
                                 // Set value with follow val from above 
                                 #tempReturnVal := "LKinLang_SetValue"(parameterValue := #tempParameterValue,
                                                                       parameterPriority := #statParameterDefinition.priorities.valueFlags.remainingDistance,
                                                                       validCountOfParameter := #statValidCounts.valueFlags.remainingDistance,
                                                                       parameterValueMin := #MINVAL_LREAL,
                                                                       parameterValueMax := #MAXVAL_LREAL,
                                                                       properties := #statParameterDefinition.properties,
                                                                       errorString => #statErrorString,
                                                                       parameterCounter := #statElementCounter.valueFlags.remainingDistance,
                                                                       priorityCounter := #statActualCommand.priority.valueFlags[#statActualValueFlagNumber].remainingDistance,
                                                                       modalCMDPrio := #statModalCommand.priority.valueFlags[#statActualValueFlagNumber].remainingDistance,
                                                                       modalPRGPrio := #statModalProgram.priority.valueFlags[#statActualValueFlagNumber].remainingDistance,
                                                                       parameterCounterInLine := #statElementCounterInLine.valueFlags.remainingDistance,
                                                                       pathDataValue := #statPathDataValue,
                                                                       modalCMDPathDataValue := #statModalCmdValue,
                                                                       modalPRGPathDataValue := #statModalPrgValue);

                                 IF #tempReturnVal = 0 THEN // Parameter is ok
                                   #statActualCommand.pathDataElement.valueFlags[#statActualValueFlagNumber].remainingDistance := #statPathDataValue.valueLReal;
                                   #statModalCommand.pathDataElement.valueFlags[#statActualValueFlagNumber].remainingDistance := #statModalCmdValue.valueLReal;
                                   #statModalProgram.pathDataElement.valueFlags[#statActualValueFlagNumber].remainingDistance := #statModalPrgValue.valueLReal;
                                 ELSE
                                   // Error
                                   #statStatus := #ERR_PARSING;
                                   #statErrorString := CONCAT(IN1 := #statErrorString, IN2 := '; Line: ');
                                   #statErrorString := CONCAT(IN1 := #statErrorString, IN2 := UDINT_TO_STRING(#statTokenizedLine.lineNo));
                                   EXIT;
                                 END_IF;
                               END_IF;

                             END_FOR;
                           END_REGION LREAL_FLAGS

                           // Exit loop in case of error
                           IF #statStatus.%X15 THEN
                             EXIT;
                           END_IF;

                         END_IF;
                       END_REGION SET_VALUES_IN_PATH_DATA_ELEMENT

                     END_FOR;

                     // Exit loop in case of error
                     IF #statStatus.%X15 THEN
                       EXIT;
                     END_IF;

                     // Check if right side of equation; if not reset it 
                     IF #statRightSideOfEquation THEN
                       ;
                     ELSE
                       #statRightSideOfEquation := TRUE;
                       #statStringExpression := '';
                     END_IF;

                     // Go to next state
                     #statStateIntern := #STATE_TOKEN_PROCESSED;

                   END_IF;
                 END_REGION TOKEN_IS_PARAMETER

                 // ------------------------------------------------------------------------------------------
                 // Is token variable
                 // Check if token is a defined variable or interface variable
                 // YES: Go to TOKEN_IS_VARIABLE
                 // NO: Go to TOKEN_IS_UNKNOWN
                 // ------------------------------------------------------------------------------------------ 
                 REGION IS_TOKEN_VARIABLE
                   IF #statStateIntern = #STATE_IS_TOKEN_VARIABLE THEN
                     // Check if token is a local or interface variable 
                     "LKinLang_IsTokenVariable"(lineNumber := #statTokenizedLine.lineNo,
                                                tokenCheck := #statTokenCheck,
                                                varIndex => #tempVarIndex,
                                                varType => #tempVarType,
                                                varRefList := #statVarRefList,
                                                keyToken := #statKeyToken,
                                                subPrgList := #statSubPrgList,
                                                errorString := #statErrorString,
                                                stringExpression := #statStringExpression);

                     // Decide where to go next
                     IF #statErrorString <> '' THEN
                       // Error occured
                       #statStateIntern := #STATE_ERROR;
                       #statStatus := #ERR_PARSING;
                       EXIT;
                     ELSIF #tempVarIndex <> 0 OR #tempVarType <> 0 THEN
                       // Go to "TOKEN_IS_VARIABLE"
                       #statStateIntern := #STATE_TOKEN_IS_VARIABLE;
                     ELSE
                       // Go to "TOKEN_IS_UNKNOWN"
                       #statStateIntern := #STATE_TOKEN_IS_UNKNOWN;
                     END_IF;
                   END_IF;
                 END_REGION IS_TOKEN_VARIABLE

                 // ------------------------------------------------------------------------------------------
                 // Token is a variable
                 // Token was found to be a valid variable
                 // SET or GET value of variable depending on context
                 // ------------------------------------------------------------------------------------------ 
                 REGION TOKEN_IS_VARIABLE
                   IF #statStateIntern = #STATE_TOKEN_IS_VARIABLE
                   THEN
                     // Token is variable 
                     // Decide if value of variable has to be set or value must be read

                     // Get value of var in following case:
                     // G0 X=myVar_1
                     // --> Variable value has to be used for X
                     // --> Concat the value to the string expression ?
                     // --> Variable is on right side of equation 
                     // Token:
                     // [1] myVar_1
                     // [2] =
                     // [3] X
                     // [4]  
                     // [5] 0
                     // [6] G

                     // Set the value of a var in following case:
                     // myVar_1 = 10 
                     // --> Variable value has to be updated
                     // --> Variable is on left side of equation
                     // 
                     // Token:
                     // [1] 10
                     // [2]
                     // [3] = 
                     // [4] 
                     // [5] myVar_1


                     IF #statRightSideOfEquation THEN
                       // --------------------------------------------------------------
                       // Right side of equation 
                       // --> GET value of variable
                       // Concat to string expression
                       // --------------------------------------------------------------
                       // Check if allowed to add number to stringExpression
                       IF "LKinLang_CharacterIsNumeric"(#statStringExpression[1]) THEN
                         // ERROR: First char is a number --> Cannot concat two numbers in a row --> ERROR
                         #statStatus := #ERR_PARSING;
                         #statErrorString := CONCAT(IN1 := #statErrorString, IN2 := 'Error: Invalid syntax');
                         #statErrorString := CONCAT(IN1 := #statErrorString, IN2 := '; Line: ');
                         #statErrorString := CONCAT(IN1 := #statErrorString, IN2 := UDINT_TO_STRING(#statTokenizedLine.lineNo));
                         EXIT;
                       ELSE
                         "LKinLang_GetVariable"(varIndex := #tempVarIndex,
                                                varType := #tempVarType,
                                                localVariables := #statVariables,
                                                interfaceVariables := #interfaceVariables,
                                                stringExpression := #statStringExpression);
                       END_IF;
                     ELSE
                       // --------------------------------------------------------------
                       // Left side of equation 
                       // --> SET value of variable
                       // Check correct syntax
                       // --------------------------------------------------------------
                       // Check if var is interface var
                       IF #tempVarType >= "LKINLANG_VAR_TYPE_INTERFACE_BOOL" THEN
                         // Previous token was index of interface var 
                         // To check correct syntax, use token before prevoius token (last but one)
                         // This token must then be a " " or "="
                         #statTokenCheck.previous := #statTokenizedLine.lineToken[#tempTokenCounter - 2];
                       END_IF;

                       // Allowed signs befor user variable
                       IF (#statTokenCheck.previous = ' '
                         XOR #statTokenCheck.previous = '=')
                       THEN // single number without _  
                         // OK
                         ;
                       ELSE
                         #statStatus := #ERR_PARSING;
                         #statStateIntern := #STATE_ERROR;
                         #statErrorString := CONCAT(IN1 := #statErrorString, IN2 := 'Error: Variable assignment');
                         #statErrorString := CONCAT(IN1 := #statErrorString, IN2 := ' in line: ');
                         #statErrorString := CONCAT(IN1 := #statErrorString, IN2 := UDINT_TO_STRING(#statTokenizedLine.lineNo));
                         EXIT;
                       END_IF;

                       // Check if variable is used a counter in for loop --> not allowed to change
                       FOR #tempCounter := 1 TO #statStack.numberOfElements DO
                         IF #statStack.stackElements[#tempCounter].variableRef.type = #tempVarType
                           AND #statStack.stackElements[#tempCounter].variableRef.index = #tempVarIndex
                         THEN
                           #statStatus := #ERR_PARSING;
                           #statStateIntern := #STATE_ERROR;
                           #statErrorString := CONCAT(IN1 := #statErrorString, IN2 := 'Error: Not allowed to change counter variable of FOR loop');
                           #statErrorString := CONCAT(IN1 := #statErrorString, IN2 := ' in line: ');
                           #statErrorString := CONCAT(IN1 := #statErrorString, IN2 := UDINT_TO_STRING(#statTokenizedLine.lineNo));
                           EXIT;
                         ELSE
                           CONTINUE;
                         END_IF;
                       END_FOR;


                       // Parse string expression and assign resulting value to variable
                       "LKinLang_SetVariable"(varIndex := #tempVarIndex,
                                              varType := #tempVarType,
                                              lineNumber := #statTokenizedLine.lineNo,
                                              stringExpression := #statStringExpression,
                                              localVariables := #statVariables,
                                              interfaceVariables := #interfaceVariables,
                                              errorString := #statErrorString);

                       IF #statErrorString <> '' THEN
                         #statStatus := #ERR_PARSING;
                         #statStateIntern := #STATE_ERROR;
                         EXIT;
                       END_IF;

                       // FR 19.03.2020
                       // Check if another assignment follows --> Keep string expression
                       IF #tempTokenCounter + 1 < #statTokenizedLine.numberOfToken THEN
                         IF #statTokenizedLine.lineToken[#tempTokenCounter + 1] <> '='
                           AND #statTokenizedLine.lineToken[#tempTokenCounter + 2] <> '=' THEN
                           // stringExpression processed --> Delete string expression
                           #statStringExpression := '';
                         END_IF;
                       ELSE
                         // stringExpression processed --> Delete string expression
                         #statStringExpression := '';
                       END_IF;

                     END_IF;

                     // Next state --> Token is processed
                     #statStateIntern := #STATE_TOKEN_PROCESSED;
                   END_IF;
                 END_REGION TOKEN_IS_VARIABLE

                 // ------------------------------------------------------------------------------------------
                 // Token is unknown
                 // Token is not a parameter or a separator 
                 // Check if equation is active and add token to string expression 
                 // If token consists of letters, it is a unknown parameter and a error is thrown
                 // Always go to TOKEN_PROCESSED
                 // ------------------------------------------------------------------------------------------ 
                 REGION TOKEN_IS_UNKNOWN
                   IF #statStateIntern = #STATE_TOKEN_IS_UNKNOWN
                   THEN

                     // Token isn't parameter
                     // Check if left side of equation
                     IF #statRightSideOfEquation = FALSE THEN
                       REGION LEFT_SIDE_EQUATION
                         // Left side of equation and no parameter 
                         // Parameter value would be handled in GetValue function in region Config commands
                         // Normally would create user variable but not implemented in V1.0
                         // Correct behaviour?
                         // Always error or concat to StringExpression ?
                         // --> Concat for something like X1=100 (More kinematics in one program)

                         // Check if token is not a number and not SPACE
                         // If yes then must be an unknwon parameter --> Error
                         IF "LKinLang_IsTokenNumber"(#statTokenCheck.actual)
                           OR "LKinLang_IsTokenNumberInclSign"(#statTokenCheck.actual)
                         THEN
                           #statStringExpression := CONCAT(IN1 := #statTokenCheck.actual, IN2 := #statStringExpression);
                         ELSE
                           // Unknon parameter
                           #statStatus := #ERR_PARSING;
                           #statErrorString := CONCAT(IN1 := #statErrorString, IN2 := 'Error unknown parameter: ');
                           #statErrorString := CONCAT(IN1 := #statErrorString, IN2 := #statTokenCheck.actual);
                           #statErrorString := CONCAT(IN1 := #statErrorString, IN2 := #statTokenCheck.previous);
                           #statErrorString := CONCAT(IN1 := #statErrorString, IN2 := '; Line: ');
                           #statErrorString := CONCAT(IN1 := #statErrorString, IN2 := UDINT_TO_STRING(#statTokenizedLine.lineNo));
                           EXIT;
                         END_IF;
                       END_REGION LEFT_SIDE_EQUATION
                     ELSE
                       REGION RIGHT_SIDE_EQUATION
                         // Token isn't parameter and right side of equation
                         // Can be a number or unknown parameter 

                         // 17.07.2019 FR: Added new check
                         // Check if token is a number
                         // Check if token is a math expression 
                         // If token is not a math expression or number then error "unknown parameter"?
                         IF "LKinLang_IsTokenNumber"(#statTokenCheck.actual)
                           OR "LKinLang_IsTokenNumberInclSign"(#statTokenCheck.actual)
                           OR "LKinLang_IsTokenMath"(#statTokenCheck.actual)
                           OR #statTokenCheck.actual = 'TRUE'
                           OR #statTokenCheck.actual = 'FALSE'
                         THEN
                           #statStringExpression := CONCAT(IN1 := #statTokenCheck.actual, IN2 := #statStringExpression);
                         ELSE
                           // Unknon parameter
                           #statStatus := #ERR_PARSING;
                           #statErrorString := CONCAT(IN1 := #statErrorString, IN2 := 'Error unknown parameter: ');
                           #statErrorString := CONCAT(IN1 := #statErrorString, IN2 := #statTokenCheck.actual);
                           #statErrorString := CONCAT(IN1 := #statErrorString, IN2 := #statTokenCheck.previous);
                           #statErrorString := CONCAT(IN1 := #statErrorString, IN2 := '; Line: ');
                           #statErrorString := CONCAT(IN1 := #statErrorString, IN2 := UDINT_TO_STRING(#statTokenizedLine.lineNo));
                           EXIT;
                         END_IF;

                       END_REGION RIGHT_SIDE_EQUATION
                     END_IF;

                     // Token is done 
                     // Go to last state
                     #statStateIntern := #STATE_TOKEN_PROCESSED;

                   END_IF;
                 END_REGION TOKEN_IS_UNKNOWN

                 // ------------------------------------------------------------------------------------------
                 // Token processed
                 // Always last state for every loop
                 // Increase token counter and check if more token follow
                 // YES: Goto STATE_INIT_PARSE_LOOP (Parse next token)
                 // NO: Goto STATE_LINE_PARSED (Line is finished)
                 // ------------------------------------------------------------------------------------------ 
                 REGION TOKEN_PROCESSED
                   // Token was processed 
                   // This is always the last state
                   IF #statStateIntern = #STATE_TOKEN_PROCESSED
                   THEN
                     #tempTokenCounter += 1;
                     IF #tempTokenCounter <= #statTokenizedLine.numberOfToken THEN
                       #statStateIntern := #STATE_INIT_PARSE_LOOP;
                     ELSE
                       #statStateIntern := #STATE_LINE_PARSED;
                     END_IF;
                   END_IF;
                 END_REGION TOKEN_PROCESSED

               END_WHILE;

             END_REGION PARSE_LINE_TOKEN

             // After the loop, check if error was set 
             IF #statStatus.%X15 THEN
               #statStateIntern := #STATE_ERROR;
             END_IF;

             // ------------------------------------------------------------------------------------------
             // Line parsed
             // Line was parsed successfully
             // Check conditions in line
             // Go to CHECK_END
             // ------------------------------------------------------------------------------------------ 
             REGION LINE_PARSED
               IF #statStateIntern = #STATE_LINE_PARSED
               THEN
                 // FR 19.03.2020:
                 // Check for missing assignment --> String expression not empty
                 IF #statStringExpression <> '' THEN
                   #statStatus := #ERR_PARSING;
                   #statStateIntern := #STATE_ERROR;
                   #statErrorString := 'Missing value assignment in line: ';
                   #statErrorString := CONCAT(IN1 := #statErrorString, IN2 := UDINT_TO_STRING(#statTokenizedLine.lineNo));

                   // Check parameter conditions in line
                 ELSIF NOT "LKinLang_CheckParameterCondition"(mode := "LKINLANG_CONDITION_IN_LINE",
                                                                language := #language,
                                                                errorString => #statErrorString,
                                                                setParameters := #statSetParametersInLine,
                                                                conditionsToCheck := #statConditionsToCheck,
                                                                parameterDefaults := #parameterDefaults)
                 THEN
                   #statStatus := #ERR_PARSING;
                   #statStateIntern := #STATE_ERROR;
                   #statErrorString := CONCAT(IN1 := #statErrorString, IN2 := ' in line: ');
                   #statErrorString := CONCAT(IN1 := #statErrorString, IN2 := UDINT_TO_STRING(#statTokenizedLine.lineNo));
                 END_IF;

                 // Go to check end
                 #statStateIntern := #STATE_CHECK_END;
               END_IF;
             END_REGION LINE_PARSED


             // ------------------------------------------------------------------------------------------
             // Check End
             // Check parsed command if cmdType = -1
             // If yes then end of program is reached and go to WRITE_COMMAND state
             // If no go to CHECK_FOR_NEW_PATH_DATA_CMD
             // ------------------------------------------------------------------------------------------ 
             REGION CHECK_END
               // Check for end of program; defined with cmdType = -1
               IF #statStateIntern = #STATE_CHECK_END
               THEN
                 IF #statActualCommand.pathDataElement.cmdType = -1
                   AND #statActualCommand.priority.cmdType > "LKINLANG_PRIO_UNRELEVANT"
                 THEN // Check for End of PRG
                   // Set execution finished if end of program is reached
                   // Status is set after command is written
                   // #statStatus := #STATUS_EXECUTION_FINISHED;

                   // Write last command with empty path data element
                   #statActualCommand.pathDataElement := #statPathDataElementEmpty.pathDataElement;

                   // Go to write command state
                   IF #statSyntaxCheck = "LKINLANG_SYNTAX_CHECK_OFF" THEN
                     #statStateIntern := #STATE_WRITE_CMD;
                     IF #lineBuffer.pointers.endOfFile = FALSE THEN
                       #lineBuffer.pointers.endOfFile := TRUE; // Signalize end to filehandler
                     END_IF;
                   ELSE
                     #statStateIntern := #STATE_RESET_AFTER_WRITE;
                   END_IF;
                   // Go to end of FOR LOOP
                   EXIT;
                 ELSE
                   // Next step --> Check if path data command is finished
                   #statStateIntern := #STATE_CHECK_FOR_NEW_PATH_DATA_CMD;
                 END_IF;
               END_IF;
             END_REGION CHECK_END

             // ------------------------------------------------------------------------------------------
             // Check for new PathDataCmd
             // End was not reached then check if parsed command is a complete PathData command
             // If yes go to state BUILD_PATH_DATA_CMD
             // If no go back to STATE_TOKENIZING (continue with next line)
             // ------------------------------------------------------------------------------------------ 
             REGION CHECK_FOR_NEW_PATH_DATA_CMD
               IF #statStateIntern = #STATE_CHECK_FOR_NEW_PATH_DATA_CMD
               THEN
                 // Check for Flag only 
                 // Flag was set but no position was programmed in the same line
                 IF ((#statActualCommand.pathDataElement.setFlags <> #statPathDataElementEmpty.pathDataElement.setFlags)
                   OR (#statActualCommand.pathDataElement.valueFlags <> #statPathDataElementEmpty.pathDataElement.valueFlags))
                   AND (#statActualCommand.priority.cmdCoordinates.cartesianPosition.x = "LKINLANG_PRIO_UNRELEVANT")
                   AND (#statActualCommand.priority.cmdCoordinates.cartesianPosition.y = "LKINLANG_PRIO_UNRELEVANT")
                   AND (#statActualCommand.priority.cmdCoordinates.cartesianPosition.z = "LKINLANG_PRIO_UNRELEVANT")
                   AND (#statActualCommand.priority.cmdCoordinates.cartesianPosition.a = "LKINLANG_PRIO_UNRELEVANT")
                   AND (#statActualCommand.priority.cmdParameters.circleParameters.auxPoint[1] = "LKINLANG_PRIO_UNRELEVANT")
                   AND (#statActualCommand.priority.cmdParameters.circleParameters.auxPoint[2] = "LKINLANG_PRIO_UNRELEVANT")
                   AND (#statActualCommand.priority.cmdParameters.circleParameters.auxPoint[3] = "LKINLANG_PRIO_UNRELEVANT")
                 THEN
                   // Flag only
                   #tempFlagOnly := TRUE;
                   // Next step --> Write PathData command to PathData
                   #statStateIntern := #STATE_BUILD_PATH_DATA_CMD;
                 ELSE

                   // Copy actual command to temp for testing if new command must be written
                   #tempTestCommand := #statActualCommand;

                   // If no motion command was parsed then use old modal command 
                   IF #tempTestCommand.motionCmd = #statPathDataElementEmpty.motionCmd THEN
                     "LKinLang_UpdateModalData"(inputPathData := #statModalCommandOld,
                                                updatedPathData := #tempTestCommand);
                   END_IF;

                   // Build complete path data command
                   // First copy CMD Modal actual command (where needed)
                   "LKinLang_UpdateModalData"(inputPathData := #statModalCommand,
                                              updatedPathData := #tempTestCommand);

                   // Second copy PRG Modal to actual command (where needed)
                   "LKinLang_UpdateModalData"(inputPathData := #statModalProgram,
                                              updatedPathData := #tempTestCommand);

                   // Check if new coordinates are set --> New path data command

                   // Testing if no cmdType is set, which one to take ?
                   IF #tempTestCommand.pathDataElement.cmdType = #statPathDataElementEmpty.pathDataElement.cmdType THEN
                     // 16.07.2019 FR: Added check of cmdType
                     // Do not always copy cmd type because LKinLang_IsNewCommand returns true if not a motion command (40,41,42, etc.)
                     IF #statActualCommandOld.pathDataElement.cmdType >= -1
                       AND #statActualCommandOld.pathDataElement.cmdType <= 4
                     THEN
                       #tempTestCommand.pathDataElement.cmdType := #statActualCommandOld.pathDataElement.cmdType;
                     END_IF;
                   END_IF;

                   IF "LKinLang_IsNewCommand"(actualPathData := #tempTestCommand,
                                                emptyPathData := #statPathDataElementEmpty,
                                                positioningMode := #statPositioningMode)
                   THEN
                     // Next step --> Write PathData command to PathData
                     #statStateIntern := #STATE_BUILD_PATH_DATA_CMD;
                   ELSE
                     // Incomplete PathData command --> Parse next line or search line
                     IF #statSearchedLine <= 0 THEN
                       // Next state --> Tokenize new line
                       #statStateIntern := #STATE_TOKENIZING;
                     ELSE
                       // Next state --> Search line
                       #statStateIntern := #STATE_SEARCH_LINE;
                     END_IF;
                   END_IF;
                 END_IF;
               END_IF;
             END_REGION CHECK_FOR_NEW_PATH_DATA_CMD

             // ------------------------------------------------------------------------------------------
             // Build PathDataCmd
             // Build complete PathData command with modal data
             // Check if all conditions are met
             // If everything is ok go to WRITE_COMMAND
             // If not go to ERROR_STATE
             // ------------------------------------------------------------------------------------------ 
             REGION BUILD_PATH_DATA_CMD
               IF #statStateIntern = #STATE_BUILD_PATH_DATA_CMD
               THEN

                 IF NOT #tempFlagOnly THEN // Normal command routine

                   REGION GET_MODAL_DATA
                     // Check if no command modal motion cmd was set; if yes assume old motion command
                     IF #statModalCommand.motionCmd = #statPathDataElementEmpty.motionCmd THEN
                       #statModalCommand.motionCmd := #statModalCommandOld.motionCmd;
                     END_IF;

                     // Update actual Command with Modal Values
                     // Check if new motion Cmd was programmed; if yes overwrite old modal cmd
                     IF #statModalCommand.motionCmd <> #statModalCommandOld.motionCmd THEN
                       // Overwrite all Old values
                       #statModalCommandOld := #statModalCommand;
                     ELSE
                       // only update values where missing
                       "LKinLang_UpdateModalData"(inputPathData := #statModalCommandOld,
                                                  updatedPathData := #statModalCommand);

                     END_IF;
                     // First copy CMD Modal to actual command (where needed)
                     "LKinLang_UpdateModalData"(inputPathData := #statModalCommand,
                                                updatedPathData := #statActualCommand);

                     // Second copy PRG Modal to actual command (where needed)
                     "LKinLang_UpdateModalData"(inputPathData := #statModalProgram,
                                                updatedPathData := #statActualCommand);

                     // --> CMD finished --> Write to PathData
                   END_REGION GET_MODAL_DATA

                   // Testing relative positioning 19.12.2018
                   REGION REL_ABS_POSITIONING
                     IF #statPositioningMode = 2 THEN // Relative
                       CASE #statActualCommand.pathDataElement.cmdType OF
                         1, 2:  // Linear command 
                           #statActualCommand.pathDataElement.cmdType := 2;
                         3, 4: // Circular command
                           #statActualCommand.pathDataElement.cmdType := 4;
                         ELSE  // Statement section ELSE
                           #statActualCommand.pathDataElement.cmdType := #statActualCommand.pathDataElement.cmdType;
                       END_CASE;

                     ELSIF #statPositioningMode = 1 THEN // Absolute
                       CASE #statActualCommand.pathDataElement.cmdType OF
                         1, 2:  // Linear command 
                           #statActualCommand.pathDataElement.cmdType := 1;
                         3, 4: // Circular command
                           #statActualCommand.pathDataElement.cmdType := 3;
                         ELSE  // Statement section ELSE
                           #statActualCommand.pathDataElement.cmdType := #statActualCommand.pathDataElement.cmdType;
                       END_CASE;
                     ELSE
                       ; // Error ?
                     END_IF;
                   END_REGION REL_ABS_POSITIONING

                 ELSE
                   // Flag only command
                   #statActualCommand.pathDataElement.cmdType := 0;
                   // Set positions zero
                   #statActualCommand.pathDataElement.cmdCoordinates.cartesianPosition.x := 0.0;
                   #statActualCommand.pathDataElement.cmdCoordinates.cartesianPosition.y := 0.0;
                   #statActualCommand.pathDataElement.cmdCoordinates.cartesianPosition.z := 0.0;
                   #statActualCommand.pathDataElement.cmdCoordinates.cartesianPosition.a := 0.0;
                   // Set all valid bits to false
                   #statActualCommand.pathDataElement.parameterValid[1] := FALSE;
                   #statActualCommand.pathDataElement.parameterValid[2] := FALSE;
                   #statActualCommand.pathDataElement.parameterValid[3] := FALSE;
                   #statActualCommand.pathDataElement.parameterValid[4] := FALSE;

                 END_IF;

                 REGION CHECK_CONDITIONS
                   // Check if conditions are met (e.g F was programmed once for G1)
                   // Check conditions in command
                   IF NOT "LKinLang_CheckParameterCondition"(mode := "LKINLANG_CONDITION_IN_COMMAND",
                                                               language := #statSelectedLanguage,
                                                               errorString => #statErrorString,
                                                               setParameters := #statSetParametersInCmd,
                                                               conditionsToCheck := #statConditionsToCheck,
                                                               parameterDefaults := #parameterDefaults)

                   THEN
                     #statStatus := #ERR_PARSING;
                     #statStateIntern := #STATE_ERROR;
                     #statErrorString := CONCAT(IN1 := #statErrorString, IN2 := ' in line: ');
                     #statErrorString := CONCAT(IN1 := #statErrorString, IN2 := UDINT_TO_STRING(#statTokenizedLine.lineNo));
                   END_IF;

                   // Check conditions in program
                   IF NOT "LKinLang_CheckParameterCondition"(mode := "LKINLANG_CONDITION_IN_PROGRAM",
                                                               language := #statSelectedLanguage,
                                                               errorString => #statErrorString,
                                                               setParameters := #statSetParametersInPrg,
                                                               conditionsToCheck := #statConditionsToCheck,
                                                               parameterDefaults := #parameterDefaults)
                   THEN
                     #statStatus := #ERR_PARSING;
                     #statStateIntern := #STATE_ERROR;
                     #statErrorString := CONCAT(IN1 := #statErrorString, IN2 := ' in line: ');
                     #statErrorString := CONCAT(IN1 := #statErrorString, IN2 := UDINT_TO_STRING(#statTokenizedLine.lineNo));
                   END_IF;
                 END_REGION CHECK_CONDITIONS

                 // Check if a flag mode was set in line
                 // If not then check the input defaults
                 // If still not set then use internal constant
                 REGION DEFAULT_FLAG_MODE

                   FOR #tempCounter := 1 TO "LKINCTRL_NO_OF_CMD_SETFLAGS" DO
                     IF #statActualCommand.pathDataElement.setFlags[#tempCounter].flag <> -1
                       AND #statActualCommand.pathDataElement.setFlags[#tempCounter].flagMode = #statParameterDefinitionEmpty.directValues.setFlags[#tempCounter].flagMode
                     THEN
                       // Check the DefaultFlagMode input for boolean flags 
                       IF #flagModeDefaults.setFlags[#statActualCommand.pathDataElement.setFlags[#tempCounter].flag].flagMode <> 0 THEN
                         #statActualCommand.pathDataElement.setFlags[#tempCounter].flagMode := #flagModeDefaults.setFlags[#statActualCommand.pathDataElement.setFlags[#tempCounter].flag].flagMode;
                       ELSE
                         #statActualCommand.pathDataElement.setFlags[#tempCounter].flagMode := #DEFAULT_FLAG_MODE;
                       END_IF;
                     END_IF;

                     // Check if flagMode 10 was set but no remaining distance
                     IF #statActualCommand.pathDataElement.setFlags[#tempCounter].flag <> -1
                       AND #statActualCommand.pathDataElement.setFlags[#tempCounter].flagMode = 10
                       AND #statActualCommand.pathDataElement.setFlags[#tempCounter].remainingDistance = #statParameterDefinitionEmpty.directValues.setFlags[#tempCounter].remainingDistance
                     THEN
                       // Check the default remainingDistance input for boolean flags 
                       IF #flagModeDefaults.setFlags[#statActualCommand.pathDataElement.setFlags[#tempCounter].flag].remainingDistance <> 0.0 THEN
                         #statActualCommand.pathDataElement.setFlags[#tempCounter].remainingDistance := #flagModeDefaults.setFlags[#statActualCommand.pathDataElement.setFlags[#tempCounter].flag].remainingDistance;
                       END_IF;
                     END_IF;
                   END_FOR;

                   FOR #tempCounter := 1 TO "LKINCTRL_NO_OF_CMD_VALUEFLAGS" DO
                     IF #statActualCommand.pathDataElement.valueFlags[#tempCounter].flag <> -1
                       AND #statActualCommand.pathDataElement.valueFlags[#tempCounter].flagMode = #statParameterDefinitionEmpty.directValues.valueFlags[#tempCounter].flagMode
                     THEN
                       // Check the DefaultFlagMode input for value flags
                       IF #flagModeDefaults.valueFlags[#statActualCommand.pathDataElement.valueFlags[#tempCounter].flag].flagMode <> 0 THEN
                         #statActualCommand.pathDataElement.valueFlags[#tempCounter].flagMode := #flagModeDefaults.valueFlags[#statActualCommand.pathDataElement.valueFlags[#tempCounter].flag].flagMode;
                       ELSE
                         #statActualCommand.pathDataElement.valueFlags[#tempCounter].flagMode := #DEFAULT_FLAG_MODE;
                       END_IF;
                     END_IF;

                     // Check if flagMode 10 was set but no remaining distance
                     IF #statActualCommand.pathDataElement.valueFlags[#tempCounter].flag <> -1
                       AND #statActualCommand.pathDataElement.valueFlags[#tempCounter].flagMode = 10
                       AND #statActualCommand.pathDataElement.valueFlags[#tempCounter].remainingDistance = #statParameterDefinitionEmpty.directValues.valueFlags[#tempCounter].remainingDistance
                     THEN
                       // Check the default remainingDistance input for value flags 
                       IF #flagModeDefaults.valueFlags[#statActualCommand.pathDataElement.valueFlags[#tempCounter].flag].remainingDistance <> 0.0 THEN
                         #statActualCommand.pathDataElement.valueFlags[#tempCounter].remainingDistance := #flagModeDefaults.valueFlags[#statActualCommand.pathDataElement.valueFlags[#tempCounter].flag].remainingDistance;
                       END_IF;
                     END_IF;
                   END_FOR;
                 END_REGION DEFAULT_FLAG_MODE

                 // Check path data command if executable / no data missing
                 #tempReturnVal := "LKinLang_CheckPathDataCmd"(errorString := #statErrorString,
                                                               pathDataCmd := #statActualCommand.pathDataElement);

                 IF #tempReturnVal <> 0 THEN
                   // Error: incomplete path data command
                   #statStatus := #ERR_PARSING;
                   #statErrorString := CONCAT(IN1 := #statErrorString, IN2 := ' in Line:');
                   #statErrorString := CONCAT(IN1 := #statErrorString, IN2 := UDINT_TO_STRING(#lineBuffer.lines[#lineBuffer.pointers.retrievePointer].number));
                   #statStateIntern := #STATE_ERROR;
                   //EXIT;
                 END_IF;

                 // Check for error while building cmd
                 IF #statStateIntern <> #STATE_ERROR THEN
                   IF #statSyntaxCheck = "LKINLANG_SYNTAX_CHECK_OFF" THEN
                     #statStateIntern := #STATE_WRITE_CMD;
                   ELSE
                     #statStateIntern := #STATE_RESET_AFTER_WRITE;
                   END_IF;
                 ELSE
                   ; // internal state is error --> Do nothing and go to error
                 END_IF;

               END_IF;
             END_REGION BUILD_PATH_DATA_CMD

             // ------------------------------------------------------------------------------------------
             // Write command
             // Building cmd is finished
             // Check PathData pointers
             // Write Command to PathData and increment pointer
             // Go to RESET_AFTER_WRITE
             // ------------------------------------------------------------------------------------------ 
             REGION WRITE_COMMAND 
               // Check if writing to PathData buffer is allowed
               IF #statStateIntern = #STATE_WRITE_CMD
                 AND
                 (((#pathData.pointers.retrievePointer <= #pathData.pointers.addPointer)
                 AND NOT #pathData.pointers.addPointerRestarted
                 AND NOT (#pathData.pointers.addPointer = "LKINCTRL_NO_OF_PATHDATA_ELEMENTS_ADVANCED"
                 AND #pathData.pointers.retrievePointer <= 1))
                 OR ((#pathData.pointers.retrievePointer > #pathData.pointers.addPointer + 1)
                 AND #pathData.pointers.addPointerRestarted))
               THEN
                 // Increment PathData buffer add pointer
                 #statAddPointer += 1;

                 // Ring buffer checks of add pointer
                 IF #statAddPointer > "LKINCTRL_NO_OF_PATHDATA_ELEMENTS_ADVANCED" THEN
                   #statAddPointer := 1;
                 END_IF;

                 // Reset path data command
                 #pathData.commands[#statAddPointer] := #statPathDataElementEmpty.pathDataElement;

                 // Copy path data element to output
                 // ---------------------------------------------------------
                 #pathData.commands[#statAddPointer] := #statActualCommand.pathDataElement;
                 // ---------------------------------------------------------

                 // Increment PathData buffer add pointer AFTER(!) writing command
                 IF #pathData.pointers.addPointer >= "LKINCTRL_NO_OF_PATHDATA_ELEMENTS_ADVANCED" AND #statAddPointer = 1 THEN
                   // Write internal to output
                   #pathData.pointers.addPointer := #statAddPointer;
                   // Set the restarted bit
                   #pathData.pointers.addPointerRestarted := TRUE;
                 ELSE
                   // Write internal to output
                   #pathData.pointers.addPointer := #statAddPointer;
                 END_IF;

                 // Reset buffer locked
                 IF #pathData.pointers.addPointer > "LKINCTRL_NO_OF_START_EXECUTE_CMDS" THEN
                   #pathData.pointers.bufferLocked := false;
                 END_IF;

                 // Next state --> Tokenize new line
                 #statStateIntern := #STATE_RESET_AFTER_WRITE;

               ELSE
                 ; // Do nothing --> error state
               END_IF;
             END_REGION WRITE_COMMAND 

             // ------------------------------------------------------------------------------------------
             // Reset variables and save "old" variables here
             // Go to STATE_TOKENIZING (continue with next line)
             // ------------------------------------------------------------------------------------------ 
             REGION RESET_AFTER_WRITE
               // Last state after writing 
               IF #statStateIntern = #STATE_RESET_AFTER_WRITE THEN

                 // If cmdType = -1 then end of parsing was found --> Execution finished
                 IF #statActualCommand.pathDataElement.cmdType = -1 THEN
                   IF #statSyntaxCheck <> "LKINLANG_SYNTAX_CHECK_AND_EXECUTE" THEN
                     // Reset line buffer retrieve pointer when finished; FR: 25.11.2019
                     #lineBuffer.pointers.retrievePointer := 0;
                     #pathData.pointers.bufferLocked := false;
                     // Reset file state
                     IF #lineBuffer.info.fileState = "LKINLANG_FILE_STATE_RUNNING" THEN
                       #lineBuffer.info.fileState := "LKINLANG_FILE_STATE_IDLE";
                     END_IF;
                     #statStatus := #STATUS_EXECUTION_FINISHED;
                   ELSE
                     // --------------------------------------------------
                     // Init variables to restart parsing and writing
                     // --------------------------------------------------
                     // Check if the line number is greater the retireve Pointer --> If yes then a buffer overflow occured and restart is neccessary
                     IF #lineBuffer.lines[#lineBuffer.pointers.retrievePointer].number > #lineBuffer.pointers.retrievePointer THEN
                       #lineBuffer.pointers.restart := TRUE;
                     END_IF;
                     // Reset line buffer retrieve pointer when finished
                     #lineBuffer.pointers.retrievePointer := 0;

                     // Set syntax check to OFF
                     #statSyntaxCheck := "LKINLANG_SYNTAX_CHECK_OFF";

                     // Init empty path data element 
                     #statModalCommand := #statPathDataElementEmpty;
                     #statModalCommandOld := #statPathDataElementEmpty;
                     #statModalProgram := #statPathDataElementEmpty;
                     #statActualCommand := #statPathDataElementEmpty;
                     #statActualCommandOld := #statPathDataElementEmpty;

                     #statElementCounter := #statElementCounterEmpty;

                     // Init conditions
                     FOR #tempCounter := 1 TO "LKINLANG_NUMBER_OF_CONDITIONS" DO
                       #statConditionsToCheck[#tempCounter] := #statConditionEmpty;
                       #statSetParametersInCmd[#tempCounter] := #statConditionEmpty;
                       #statSetParametersInPrg[#tempCounter] := #statConditionEmpty;
                     END_FOR;

                     // Init tokenized line
                     #statTokenizedLine.lineNo := 0;
                     #statTokenizedLine.numberOfToken := 0;
                     FOR #tempCounter := 1 TO "LKINLANG_MAX_NUMBER_OF_TOKEN_PER_LINE" DO
                       #statTokenizedLine.lineToken[#tempCounter] := '';
                     END_FOR;

                     // Init Positioning mode to absolute
                     #statPositioningMode := 1;

                     // Init token counter
                     #tempTokenCounter := 1;

                     // Init condition counter
                     #tempConditionCounter := 1;

                     // Init flag counter
                     #statActualFlagNumber := 0;

                     // Reset varaibles to avoid duplcate errors
                     // Init vars & counter
                     FOR #tempVarIndex := 1 TO "LKINLANG_NUMBER_OF_LOCAL_BOOL" DO
                       #statVariables.boolean[#tempVarIndex] := FALSE;
                     END_FOR;
                     FOR #tempVarIndex := 1 TO "LKINLANG_NUMBER_OF_LOCAL_DINT" DO
                       #statVariables.dints[#tempVarIndex] := 0;
                     END_FOR;
                     FOR #tempVarIndex := 1 TO "LKINLANG_NUMBER_OF_LOCAL_LREAL" DO
                       #statVariables.lreals[#tempVarIndex] := 0.0;
                     END_FOR;
                     #statVariables.boolCounter := 0;
                     #statVariables.dintCounter := 0;
                     #statVariables.lrealCounter := 0;

                     // Remove local vars from var ref table
                     FOR #tempVarIndex := 1 TO "LKINLANG_NUMBER_OF_VAR_REFS" DO
                       IF #statVarRefList.references[#tempVarIndex].type < "LKINLANG_VAR_TYPE_INTERFACE_BOOL" THEN
                         #statVarRefList.references[#tempVarIndex].index := 0;
                         #statVarRefList.references[#tempVarIndex].name := '';
                         #statVarRefList.references[#tempVarIndex].type := 0;
                       END_IF;
                     END_FOR;

                     // TODO: Check if reset is OK!
                     #statVarRefList.numberOfReferences := 0;
                   END_IF;

                 END_IF;

